REGION Network 14: I42.5 - Tank Vent Valve 2 Feedback Closed (CV-441-B)
   // True = CLOSED, False = NOT
   RUNG wire#powerrail
      Contact( "Tank 4S Tank Vent Valve 2 Feedback - Closed" )
      Coil( "20_TANKS_IP_DATA".RIO_04.SECOND_TANK.TANK_VENT_B_CLSD )
   END_RUNG
   // the same network as SCL:
   "20_TANKS_IP_DATA".RIO_04.SECOND_TANK.TANK_VENT_B_CLSD := "Tank 4S Tank Vent Valve 2 Feedback - Closed";
END_REGION

REGION Network 15: I42.6 - Spare Input Destination Accesed from Warning FC
   // True = N/A, False = N/A
END_REGION

REGION Network 16: I42.7 - Spare Input
   // True = N/A, False = N/A
   RUNG wire#powerrail
      Contact( "RIO4_SPR_DI_142_7" )
      Coil( "20_TANKS_IP_DATA".RIO_04.SECOND_TANK.SPARE_DI_7 )
   END_RUNG
   // the same network as SCL:
   "20_TANKS_IP_DATA".RIO_04.SECOND_TANK.SPARE_DI_7 := "RIO4_SPR_DI_142_7";
END_REGION

REGION Network 17: I45.0 - Tank Level HIHI - (LS-425) - First Tank
   // True = OK, False = HIHI
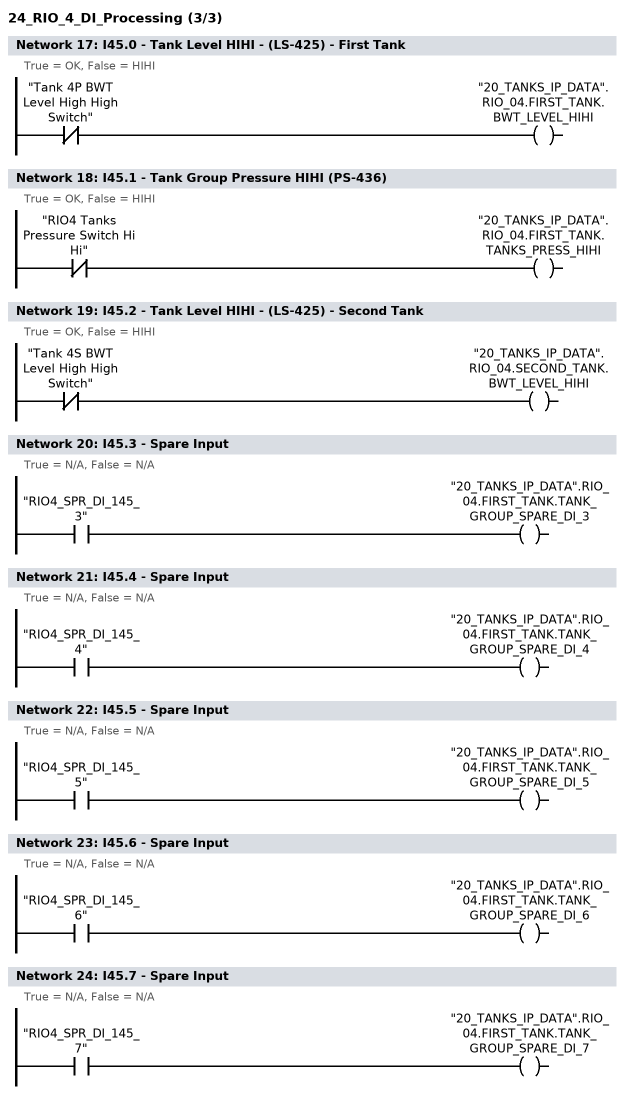
   RUNG wire#powerrail
      I_Contact( "Tank 4P BWT Level High High Switch" )
      Coil( "20_TANKS_IP_DATA".RIO_04.FIRST_TANK.BWT_LEVEL_HIHI )
   END_RUNG
   // the same network as SCL:
   "20_TANKS_IP_DATA".RIO_04.FIRST_TANK.BWT_LEVEL_HIHI := NOT "Tank 4P BWT Level High High Switch";
END_REGION

REGION Network 18: I45.1 - Tank Group Pressure HIHI (PS-436)
   // True = OK, False = HIHI
   RUNG wire#powerrail
      I_Contact( "RIO4 Tanks Pressure Switch Hi Hi" )
      Coil( "20_TANKS_IP_DATA".RIO_04.FIRST_TANK.TANKS_PRESS_HIHI )
   END_RUNG
   // the same network as SCL:
   "20_TANKS_IP_DATA".RIO_04.FIRST_TANK.TANKS_PRESS_HIHI := NOT "RIO4 Tanks Pressure Switch Hi Hi";
END_REGION

REGION Network 19: I45.2 - Tank Level HIHI - (LS-425) - Second Tank
   // True = OK, False = HIHI
   RUNG wire#powerrail
      I_Contact( "Tank 4S BWT Level High High Switch" )
      Coil( "20_TANKS_IP_DATA".RIO_04.SECOND_TANK.BWT_LEVEL_HIHI )
   END_RUNG
   // the same network as SCL:
   "20_TANKS_IP_DATA".RIO_04.SECOND_TANK.BWT_LEVEL_HIHI := NOT "Tank 4S BWT Level High High Switch";
END_REGION

REGION Network 20: I45.3 - Spare Input
   // True = N/A, False = N/A
   RUNG wire#powerrail
      Contact( "RIO4_SPR_DI_145_3" )
      Coil( "20_TANKS_IP_DATA".RIO_04.FIRST_TANK.TANK_GROUP_SPARE_DI_3 )
   END_RUNG
   // the same network as SCL:
   "20_TANKS_IP_DATA".RIO_04.FIRST_TANK.TANK_GROUP_SPARE_DI_3 := "RIO4_SPR_DI_145_3";
END_REGION

REGION Network 21: I45.4 - Spare Input
   // True = N/A, False = N/A
   RUNG wire#powerrail
      Contact( "RIO4_SPR_DI_145_4" )
      Coil( "20_TANKS_IP_DATA".RIO_04.FIRST_TANK.TANK_GROUP_SPARE_DI_4 )
   END_RUNG
   // the same network as SCL:
   "20_TANKS_IP_DATA".RIO_04.FIRST_TANK.TANK_GROUP_SPARE_DI_4 := "RIO4_SPR_DI_145_4";
END_REGION

REGION Network 22: I45.5 - Spare Input
   // True = N/A, False = N/A
   RUNG wire#powerrail
      Contact( "RIO4_SPR_DI_145_5" )
      Coil( "20_TANKS_IP_DATA".RIO_04.FIRST_TANK.TANK_GROUP_SPARE_DI_5 )
   END_RUNG
   // the same network as SCL:
   "20_TANKS_IP_DATA".RIO_04.FIRST_TANK.TANK_GROUP_SPARE_DI_5 := "RIO4_SPR_DI_145_5";
END_REGION

REGION Network 23: I45.6 - Spare Input
   // True = N/A, False = N/A
   RUNG wire#powerrail
      Contact( "RIO4_SPR_DI_145_6" )
      Coil( "20_TANKS_IP_DATA".RIO_04.FIRST_TANK.TANK_GROUP_SPARE_DI_6 )
   END_RUNG
   // the same network as SCL:
   "20_TANKS_IP_DATA".RIO_04.FIRST_TANK.TANK_GROUP_SPARE_DI_6 := "RIO4_SPR_DI_145_6";
END_REGION

REGION Network 24: I45.7 - Spare Input
   // True = N/A, False = N/A
   RUNG wire#powerrail
      Contact( "RIO4_SPR_DI_145_7" )
      Coil( "20_TANKS_IP_DATA".RIO_04.FIRST_TANK.TANK_GROUP_SPARE_DI_7 )
   END_RUNG
   // the same network as SCL:
   "20_TANKS_IP_DATA".RIO_04.FIRST_TANK.TANK_GROUP_SPARE_DI_7 := "RIO4_SPR_DI_145_7";
END_REGION
END_FUNCTION

FUNCTION "25_RIO_5_DI_Processing" : Void   // FC25, LAD
TITLE = RIO Rack Digital Input Processing (Tank 1 = 5P, Tank 2 = 5S)
{ S7_Optimized_Access := 'TRUE' }
AUTHOR : JRS
VERSION : 0.1
// To process raw inputs prior to code use
BEGIN

REGION Network 1: I51.0 - Gas To Tank Valve Feedback Open (CV-422)
   // True = OPEN, False = NOT
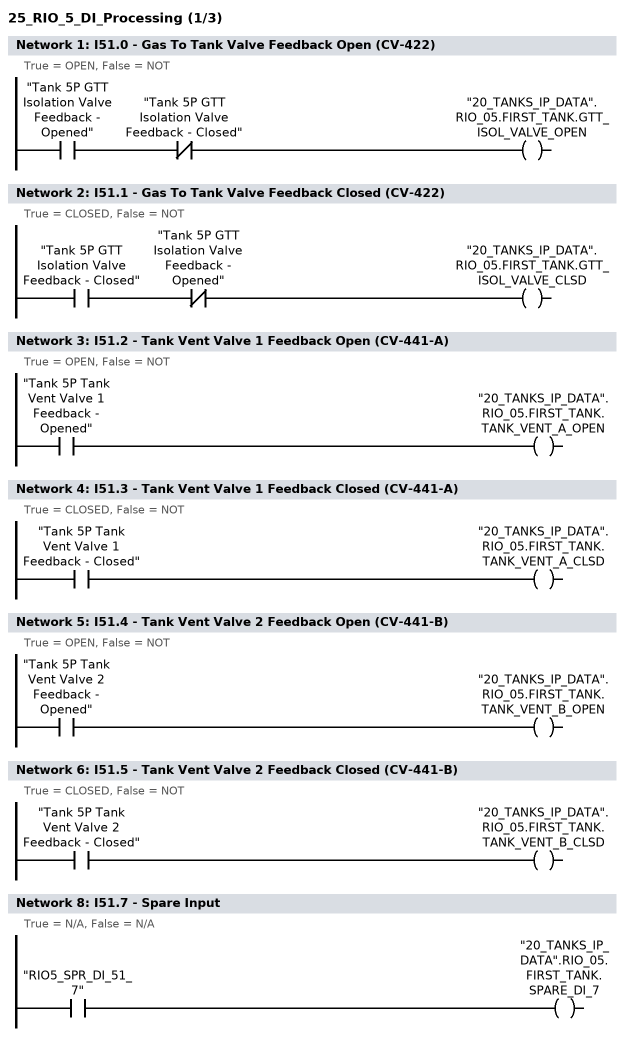
   RUNG wire#powerrail
      Contact( "Tank 5P GTT Isolation Valve Feedback - Opened" )
      I_Contact( "Tank 5P GTT Isolation Valve Feedback - Closed" )
      Coil( "20_TANKS_IP_DATA".RIO_05.FIRST_TANK.GTT_ISOL_VALVE_OPEN )
   END_RUNG
   // the same network as SCL:
   "20_TANKS_IP_DATA".RIO_05.FIRST_TANK.GTT_ISOL_VALVE_OPEN := "Tank 5P GTT Isolation Valve Feedback - Opened" AND NOT "Tank 5P GTT Isolation Valve Feedback - Closed";
END_REGION

REGION Network 2: I51.1 - Gas To Tank Valve Feedback Closed (CV-422)
   // True = CLOSED, False = NOT
   RUNG wire#powerrail
      Contact( "Tank 5P GTT Isolation Valve Feedback - Closed" )
      I_Contact( "Tank 5P GTT Isolation Valve Feedback - Opened" )
      Coil( "20_TANKS_IP_DATA".RIO_05.FIRST_TANK.GTT_ISOL_VALVE_CLSD )
   END_RUNG
   // the same network as SCL:
   "20_TANKS_IP_DATA".RIO_05.FIRST_TANK.GTT_ISOL_VALVE_CLSD := "Tank 5P GTT Isolation Valve Feedback - Closed" AND NOT "Tank 5P GTT Isolation Valve Feedback - Opened";
END_REGION

REGION Network 3: I51.2 - Tank Vent Valve 1 Feedback Open (CV-441-A)
   // True = OPEN, False = NOT
   RUNG wire#powerrail
      Contact( "Tank 5P Tank Vent Valve 1 Feedback - Opened" )
      Coil( "20_TANKS_IP_DATA".RIO_05.FIRST_TANK.TANK_VENT_A_OPEN )
   END_RUNG
   // the same network as SCL:
   "20_TANKS_IP_DATA".RIO_05.FIRST_TANK.TANK_VENT_A_OPEN := "Tank 5P Tank Vent Valve 1 Feedback - Opened";
END_REGION

REGION Network 4: I51.3 - Tank Vent Valve 1 Feedback Closed (CV-441-A)
   // True = CLOSED, False = NOT
   RUNG wire#powerrail
      Contact( "Tank 5P Tank Vent Valve 1 Feedback - Closed" )
      Coil( "20_TANKS_IP_DATA".RIO_05.FIRST_TANK.TANK_VENT_A_CLSD )
   END_RUNG
   // the same network as SCL:
   "20_TANKS_IP_DATA".RIO_05.FIRST_TANK.TANK_VENT_A_CLSD := "Tank 5P Tank Vent Valve 1 Feedback - Closed";
END_REGION

REGION Network 5: I51.4 - Tank Vent Valve 2 Feedback Open (CV-441-B)
   // True = OPEN, False = NOT
   RUNG wire#powerrail
      Contact( "Tank 5P Tank Vent Valve 2 Feedback - Opened" )
      Coil( "20_TANKS_IP_DATA".RIO_05.FIRST_TANK.TANK_VENT_B_OPEN )
   END_RUNG
   // the same network as SCL:
   "20_TANKS_IP_DATA".RIO_05.FIRST_TANK.TANK_VENT_B_OPEN := "Tank 5P Tank Vent Valve 2 Feedback - Opened";
END_REGION

REGION Network 6: I51.5 - Tank Vent Valve 2 Feedback Closed (CV-441-B)
   // True = CLOSED, False = NOT
   RUNG wire#powerrail
      Contact( "Tank 5P Tank Vent Valve 2 Feedback - Closed" )
      Coil( "20_TANKS_IP_DATA".RIO_05.FIRST_TANK.TANK_VENT_B_CLSD )
   END_RUNG
   // the same network as SCL:
   "20_TANKS_IP_DATA".RIO_05.FIRST_TANK.TANK_VENT_B_CLSD := "Tank 5P Tank Vent Valve 2 Feedback - Closed";
END_REGION

REGION Network 7: I51.6 - Spare Input Destination Accesed from Warning FC
   // True = N/A, False = N/A
END_REGION

REGION Network 8: I51.7 - Spare Input
   // True = N/A, False = N/A
   RUNG wire#powerrail
      Contact( "RIO5_SPR_DI_51_7" )
      Coil( "20_TANKS_IP_DATA".RIO_05.FIRST_TANK.SPARE_DI_7 )
   END_RUNG
   // the same network as SCL:
   "20_TANKS_IP_DATA".RIO_05.FIRST_TANK.SPARE_DI_7 := "RIO5_SPR_DI_51_7";
END_REGION

REGION Network 9: I54.0 - Gas To Tank Valve Feedback Open (CV-422)
   // True = OPEN, False = NOT
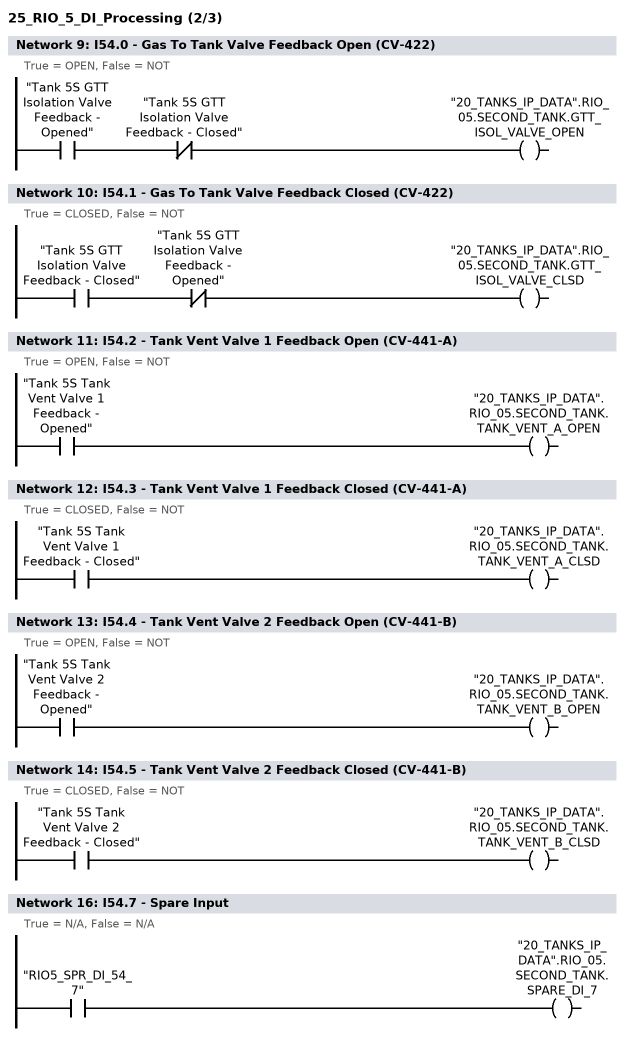
   RUNG wire#powerrail
      Contact( "Tank 5S GTT Isolation Valve Feedback - Opened" )
      I_Contact( "Tank 5S GTT Isolation Valve Feedback - Closed" )
      Coil( "20_TANKS_IP_DATA".RIO_05.SECOND_TANK.GTT_ISOL_VALVE_OPEN )
   END_RUNG
   // the same network as SCL:
   "20_TANKS_IP_DATA".RIO_05.SECOND_TANK.GTT_ISOL_VALVE_OPEN := "Tank 5S GTT Isolation Valve Feedback - Opened" AND NOT "Tank 5S GTT Isolation Valve Feedback - Closed";
END_REGION

REGION Network 10: I54.1 - Gas To Tank Valve Feedback Closed (CV-422)
   // True = CLOSED, False = NOT
   RUNG wire#powerrail
      Contact( "Tank 5S GTT Isolation Valve Feedback - Closed" )
      I_Contact( "Tank 5S GTT Isolation Valve Feedback - Opened" )
      Coil( "20_TANKS_IP_DATA".RIO_05.SECOND_TANK.GTT_ISOL_VALVE_CLSD )
   END_RUNG
   // the same network as SCL:
   "20_TANKS_IP_DATA".RIO_05.SECOND_TANK.GTT_ISOL_VALVE_CLSD := "Tank 5S GTT Isolation Valve Feedback - Closed" AND NOT "Tank 5S GTT Isolation Valve Feedback - Opened";
END_REGION

REGION Network 11: I54.2 - Tank Vent Valve 1 Feedback Open (CV-441-A)
   // True = OPEN, False = NOT
   RUNG wire#powerrail
      Contact( "Tank 5S Tank Vent Valve 1 Feedback - Opened" )
      Coil( "20_TANKS_IP_DATA".RIO_05.SECOND_TANK.TANK_VENT_A_OPEN )
   END_RUNG
   // the same network as SCL:
   "20_TANKS_IP_DATA".RIO_05.SECOND_TANK.TANK_VENT_A_OPEN := "Tank 5S Tank Vent Valve 1 Feedback - Opened";
END_REGION

REGION Network 12: I54.3 - Tank Vent Valve 1 Feedback Closed (CV-441-A)
   // True = CLOSED, False = NOT
   RUNG wire#powerrail
      Contact( "Tank 5S Tank Vent Valve 1 Feedback - Closed" )
      Coil( "20_TANKS_IP_DATA".RIO_05.SECOND_TANK.TANK_VENT_A_CLSD )
   END_RUNG
   // the same network as SCL:
   "20_TANKS_IP_DATA".RIO_05.SECOND_TANK.TANK_VENT_A_CLSD := "Tank 5S Tank Vent Valve 1 Feedback - Closed";
END_REGION

REGION Network 13: I54.4 - Tank Vent Valve 2 Feedback Open (CV-441-B)
   // True = OPEN, False = NOT
   RUNG wire#powerrail
      Contact( "Tank 5S Tank Vent Valve 2 Feedback - Opened" )
      Coil( "20_TANKS_IP_DATA".RIO_05.SECOND_TANK.TANK_VENT_B_OPEN )
   END_RUNG
   // the same network as SCL:
   "20_TANKS_IP_DATA".RIO_05.SECOND_TANK.TANK_VENT_B_OPEN := "Tank 5S Tank Vent Valve 2 Feedback - Opened";
END_REGION

REGION Network 14: I54.5 - Tank Vent Valve 2 Feedback Closed (CV-441-B)
   // True = CLOSED, False = NOT
   RUNG wire#powerrail
      Contact( "Tank 5S Tank Vent Valve 2 Feedback - Closed" )
      Coil( "20_TANKS_IP_DATA".RIO_05.SECOND_TANK.TANK_VENT_B_CLSD )
   END_RUNG
   // the same network as SCL:
   "20_TANKS_IP_DATA".RIO_05.SECOND_TANK.TANK_VENT_B_CLSD := "Tank 5S Tank Vent Valve 2 Feedback - Closed";
END_REGION

REGION Network 15: I54.6 - Spare Input Destination Accesed from Warning FC
   // True = N/A, False = N/A
END_REGION

REGION Network 16: I54.7 - Spare Input
   // True = N/A, False = N/A
   RUNG wire#powerrail
      Contact( "RIO5_SPR_DI_54_7" )
      Coil( "20_TANKS_IP_DATA".RIO_05.SECOND_TANK.SPARE_DI_7 )
   END_RUNG
   // the same network as SCL:
   "20_TANKS_IP_DATA".RIO_05.SECOND_TANK.SPARE_DI_7 := "RIO5_SPR_DI_54_7";
END_REGION

REGION Network 17: I57.0 - Tank Level HIHI - (LS-425) - First Tank
   // True = OK, False = HIHI
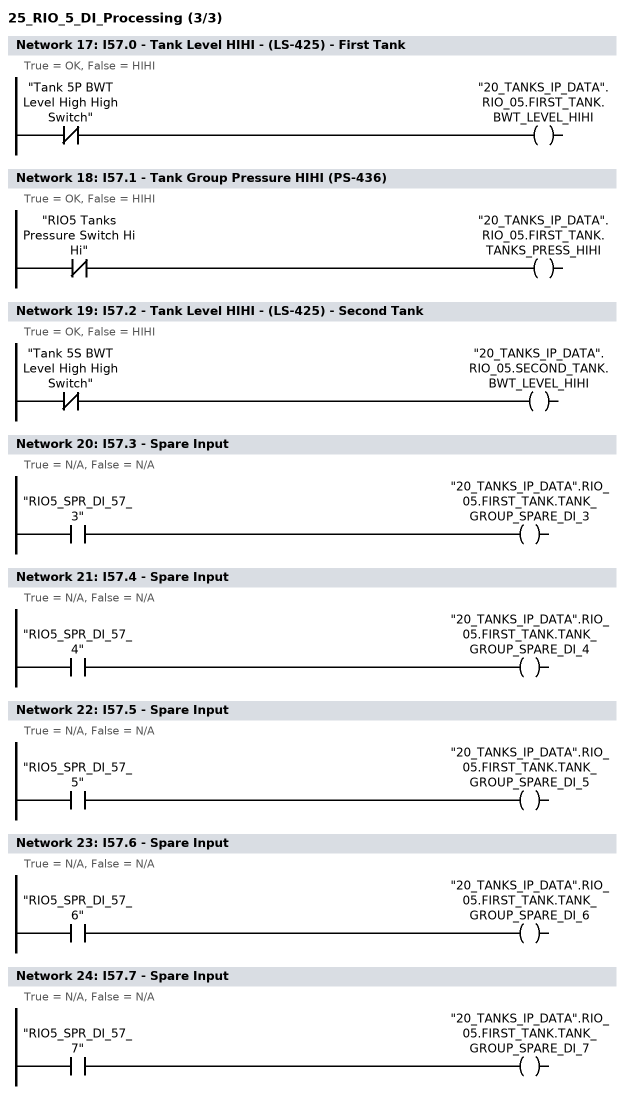
   RUNG wire#powerrail
      I_Contact( "Tank 5P BWT Level High High Switch" )
      Coil( "20_TANKS_IP_DATA".RIO_05.FIRST_TANK.BWT_LEVEL_HIHI )
   END_RUNG
   // the same network as SCL:
   "20_TANKS_IP_DATA".RIO_05.FIRST_TANK.BWT_LEVEL_HIHI := NOT "Tank 5P BWT Level High High Switch";
END_REGION

REGION Network 18: I57.1 - Tank Group Pressure HIHI (PS-436)
   // True = OK, False = HIHI
   RUNG wire#powerrail
      I_Contact( "RIO5 Tanks Pressure Switch Hi Hi" )
      Coil( "20_TANKS_IP_DATA".RIO_05.FIRST_TANK.TANKS_PRESS_HIHI )
   END_RUNG
   // the same network as SCL:
   "20_TANKS_IP_DATA".RIO_05.FIRST_TANK.TANKS_PRESS_HIHI := NOT "RIO5 Tanks Pressure Switch Hi Hi";
END_REGION

REGION Network 19: I57.2 - Tank Level HIHI - (LS-425) - Second Tank
   // True = OK, False = HIHI
   RUNG wire#powerrail
      I_Contact( "Tank 5S BWT Level High High Switch" )
      Coil( "20_TANKS_IP_DATA".RIO_05.SECOND_TANK.BWT_LEVEL_HIHI )
   END_RUNG
   // the same network as SCL:
   "20_TANKS_IP_DATA".RIO_05.SECOND_TANK.BWT_LEVEL_HIHI := NOT "Tank 5S BWT Level High High Switch";
END_REGION

REGION Network 20: I57.3 - Spare Input
   // True = N/A, False = N/A
   RUNG wire#powerrail
      Contact( "RIO5_SPR_DI_57_3" )
      Coil( "20_TANKS_IP_DATA".RIO_05.FIRST_TANK.TANK_GROUP_SPARE_DI_3 )
   END_RUNG
   // the same network as SCL:
   "20_TANKS_IP_DATA".RIO_05.FIRST_TANK.TANK_GROUP_SPARE_DI_3 := "RIO5_SPR_DI_57_3";
END_REGION

REGION Network 21: I57.4 - Spare Input
   // True = N/A, False = N/A
   RUNG wire#powerrail
      Contact( "RIO5_SPR_DI_57_4" )
      Coil( "20_TANKS_IP_DATA".RIO_05.FIRST_TANK.TANK_GROUP_SPARE_DI_4 )
   END_RUNG
   // the same network as SCL:
   "20_TANKS_IP_DATA".RIO_05.FIRST_TANK.TANK_GROUP_SPARE_DI_4 := "RIO5_SPR_DI_57_4";
END_REGION

REGION Network 22: I57.5 - Spare Input
   // True = N/A, False = N/A
   RUNG wire#powerrail
      Contact( "RIO5_SPR_DI_57_5" )
      Coil( "20_TANKS_IP_DATA".RIO_05.FIRST_TANK.TANK_GROUP_SPARE_DI_5 )
   END_RUNG
   // the same network as SCL:
   "20_TANKS_IP_DATA".RIO_05.FIRST_TANK.TANK_GROUP_SPARE_DI_5 := "RIO5_SPR_DI_57_5";
END_REGION

REGION Network 23: I57.6 - Spare Input
   // True = N/A, False = N/A
   RUNG wire#powerrail
      Contact( "RIO5_SPR_DI_57_6" )
      Coil( "20_TANKS_IP_DATA".RIO_05.FIRST_TANK.TANK_GROUP_SPARE_DI_6 )
   END_RUNG
   // the same network as SCL:
   "20_TANKS_IP_DATA".RIO_05.FIRST_TANK.TANK_GROUP_SPARE_DI_6 := "RIO5_SPR_DI_57_6";
END_REGION

REGION Network 24: I57.7 - Spare Input
   // True = N/A, False = N/A
   RUNG wire#powerrail
      Contact( "RIO5_SPR_DI_57_7" )
      Coil( "20_TANKS_IP_DATA".RIO_05.FIRST_TANK.TANK_GROUP_SPARE_DI_7 )
   END_RUNG
   // the same network as SCL:
   "20_TANKS_IP_DATA".RIO_05.FIRST_TANK.TANK_GROUP_SPARE_DI_7 := "RIO5_SPR_DI_57_7";
END_REGION
END_FUNCTION

FUNCTION "26_RIO_6_DI_Processing" : Void   // FC26, LAD
TITLE = RIO Rack Digital Input Processing (Tank 1 = 6P, Tank 2 = 6S)
{ S7_Optimized_Access := 'TRUE' }
AUTHOR : JRS
VERSION : 0.1
// To process raw inputs prior to code use
BEGIN

REGION Network 1: I60.0 - Gas To Tank Valve Feedback Open (CV-422)
   // True = OPEN, False = NOT
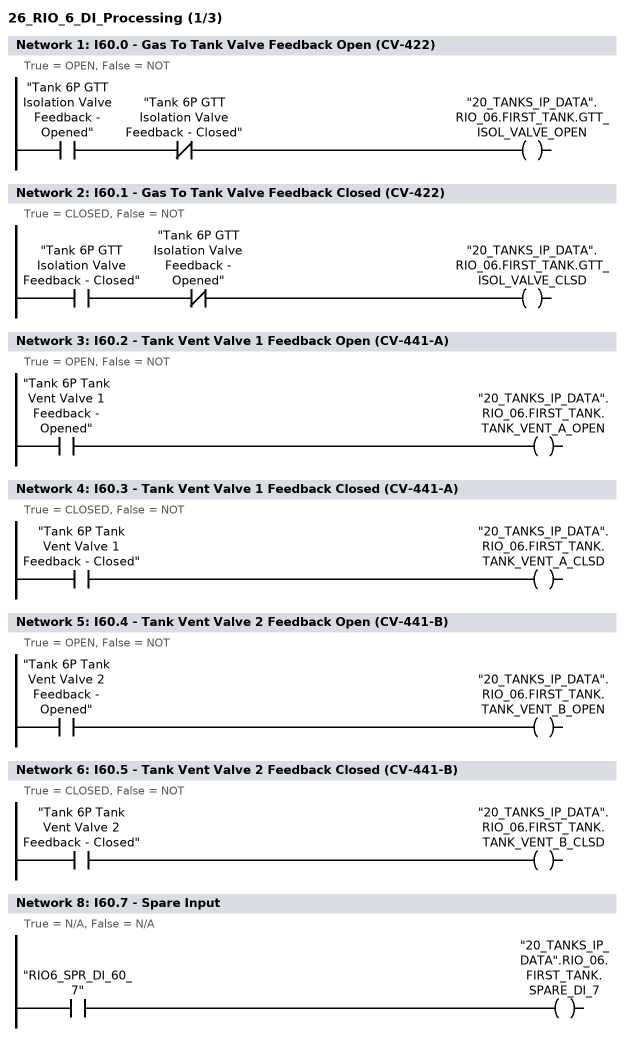
   RUNG wire#powerrail
      Contact( "Tank 6P GTT Isolation Valve Feedback - Opened" )
      I_Contact( "Tank 6P GTT Isolation Valve Feedback - Closed" )
      Coil( "20_TANKS_IP_DATA".RIO_06.FIRST_TANK.GTT_ISOL_VALVE_OPEN )
   END_RUNG
   // the same network as SCL:
   "20_TANKS_IP_DATA".RIO_06.FIRST_TANK.GTT_ISOL_VALVE_OPEN := "Tank 6P GTT Isolation Valve Feedback - Opened" AND NOT "Tank 6P GTT Isolation Valve Feedback - Closed";
END_REGION

REGION Network 2: I60.1 - Gas To Tank Valve Feedback Closed (CV-422)
   // True = CLOSED, False = NOT
   RUNG wire#powerrail
      Contact( "Tank 6P GTT Isolation Valve Feedback - Closed" )
      I_Contact( "Tank 6P GTT Isolation Valve Feedback - Opened" )
      Coil( "20_TANKS_IP_DATA".RIO_06.FIRST_TANK.GTT_ISOL_VALVE_CLSD )
   END_RUNG
   // the same network as SCL:
   "20_TANKS_IP_DATA".RIO_06.FIRST_TANK.GTT_ISOL_VALVE_CLSD := "Tank 6P GTT Isolation Valve Feedback - Closed" AND NOT "Tank 6P GTT Isolation Valve Feedback - Opened";
END_REGION

REGION Network 3: I60.2 - Tank Vent Valve 1 Feedback Open (CV-441-A)
   // True = OPEN, False = NOT
   RUNG wire#powerrail
      Contact( "Tank 6P Tank Vent Valve 1 Feedback - Opened" )
      Coil( "20_TANKS_IP_DATA".RIO_06.FIRST_TANK.TANK_VENT_A_OPEN )
   END_RUNG
   // the same network as SCL:
   "20_TANKS_IP_DATA".RIO_06.FIRST_TANK.TANK_VENT_A_OPEN := "Tank 6P Tank Vent Valve 1 Feedback - Opened";
END_REGION

REGION Network 4: I60.3 - Tank Vent Valve 1 Feedback Closed (CV-441-A)
   // True = CLOSED, False = NOT
   RUNG wire#powerrail
      Contact( "Tank 6P Tank Vent Valve 1 Feedback - Closed" )
      Coil( "20_TANKS_IP_DATA".RIO_06.FIRST_TANK.TANK_VENT_A_CLSD )
   END_RUNG
   // the same network as SCL:
   "20_TANKS_IP_DATA".RIO_06.FIRST_TANK.TANK_VENT_A_CLSD := "Tank 6P Tank Vent Valve 1 Feedback - Closed";
END_REGION

REGION Network 5: I60.4 - Tank Vent Valve 2 Feedback Open (CV-441-B)
   // True = OPEN, False = NOT
   RUNG wire#powerrail
      Contact( "Tank 6P Tank Vent Valve 2 Feedback - Opened" )
      Coil( "20_TANKS_IP_DATA".RIO_06.FIRST_TANK.TANK_VENT_B_OPEN )
   END_RUNG
   // the same network as SCL:
   "20_TANKS_IP_DATA".RIO_06.FIRST_TANK.TANK_VENT_B_OPEN := "Tank 6P Tank Vent Valve 2 Feedback - Opened";
END_REGION

REGION Network 6: I60.5 - Tank Vent Valve 2 Feedback Closed (CV-441-B)
   // True = CLOSED, False = NOT
   RUNG wire#powerrail
      Contact( "Tank 6P Tank Vent Valve 2 Feedback - Closed" )
      Coil( "20_TANKS_IP_DATA".RIO_06.FIRST_TANK.TANK_VENT_B_CLSD )
   END_RUNG
   // the same network as SCL:
   "20_TANKS_IP_DATA".RIO_06.FIRST_TANK.TANK_VENT_B_CLSD := "Tank 6P Tank Vent Valve 2 Feedback - Closed";
END_REGION

REGION Network 7: I60.6 - Spare Input Destination Accesed from Warning FC
   // True = N/A, False = N/A
END_REGION

REGION Network 8: I60.7 - Spare Input
   // True = N/A, False = N/A
   RUNG wire#powerrail
      Contact( "RIO6_SPR_DI_60_7" )
      Coil( "20_TANKS_IP_DATA".RIO_06.FIRST_TANK.SPARE_DI_7 )
   END_RUNG
   // the same network as SCL:
   "20_TANKS_IP_DATA".RIO_06.FIRST_TANK.SPARE_DI_7 := "RIO6_SPR_DI_60_7";
END_REGION

REGION Network 9: I63.0 - Gas To Tank Valve Feedback Open (CV-422)
   // True = OPEN, False = NOT
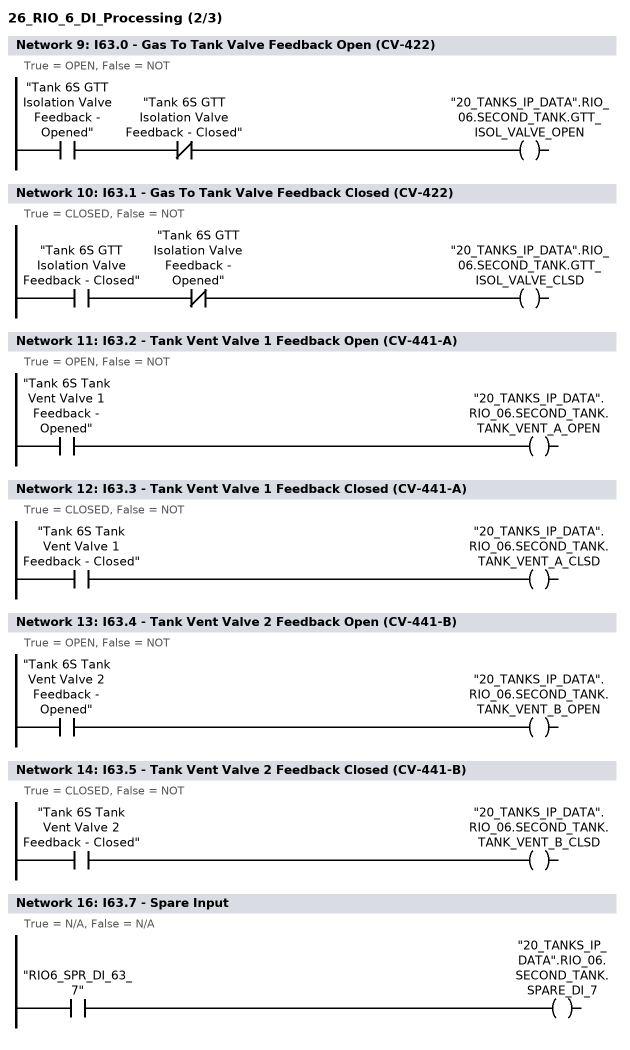
   RUNG wire#powerrail
      Contact( "Tank 6S GTT Isolation Valve Feedback - Opened" )
      I_Contact( "Tank 6S GTT Isolation Valve Feedback - Closed" )
      Coil( "20_TANKS_IP_DATA".RIO_06.SECOND_TANK.GTT_ISOL_VALVE_OPEN )
   END_RUNG
   // the same network as SCL:
   "20_TANKS_IP_DATA".RIO_06.SECOND_TANK.GTT_ISOL_VALVE_OPEN := "Tank 6S GTT Isolation Valve Feedback - Opened" AND NOT "Tank 6S GTT Isolation Valve Feedback - Closed";
END_REGION

REGION Network 10: I63.1 - Gas To Tank Valve Feedback Closed (CV-422)
   // True = CLOSED, False = NOT
   RUNG wire#powerrail
      Contact( "Tank 6S GTT Isolation Valve Feedback - Closed" )
      I_Contact( "Tank 6S GTT Isolation Valve Feedback - Opened" )
      Coil( "20_TANKS_IP_DATA".RIO_06.SECOND_TANK.GTT_ISOL_VALVE_CLSD )
   END_RUNG
   // the same network as SCL:
   "20_TANKS_IP_DATA".RIO_06.SECOND_TANK.GTT_ISOL_VALVE_CLSD := "Tank 6S GTT Isolation Valve Feedback - Closed" AND NOT "Tank 6S GTT Isolation Valve Feedback - Opened";
END_REGION

REGION Network 11: I63.2 - Tank Vent Valve 1 Feedback Open (CV-441-A)
   // True = OPEN, False = NOT
   RUNG wire#powerrail
      Contact( "Tank 6S Tank Vent Valve 1 Feedback - Opened" )
      Coil( "20_TANKS_IP_DATA".RIO_06.SECOND_TANK.TANK_VENT_A_OPEN )
   END_RUNG
   // the same network as SCL:
   "20_TANKS_IP_DATA".RIO_06.SECOND_TANK.TANK_VENT_A_OPEN := "Tank 6S Tank Vent Valve 1 Feedback - Opened";
END_REGION

REGION Network 12: I63.3 - Tank Vent Valve 1 Feedback Closed (CV-441-A)
   // True = CLOSED, False = NOT
   RUNG wire#powerrail
      Contact( "Tank 6S Tank Vent Valve 1 Feedback - Closed" )
      Coil( "20_TANKS_IP_DATA".RIO_06.SECOND_TANK.TANK_VENT_A_CLSD )
   END_RUNG
   // the same network as SCL:
   "20_TANKS_IP_DATA".RIO_06.SECOND_TANK.TANK_VENT_A_CLSD := "Tank 6S Tank Vent Valve 1 Feedback - Closed";
END_REGION

REGION Network 13: I63.4 - Tank Vent Valve 2 Feedback Open (CV-441-B)
   // True = OPEN, False = NOT
   RUNG wire#powerrail
      Contact( "Tank 6S Tank Vent Valve 2 Feedback - Opened" )
      Coil( "20_TANKS_IP_DATA".RIO_06.SECOND_TANK.TANK_VENT_B_OPEN )
   END_RUNG
   // the same network as SCL:
   "20_TANKS_IP_DATA".RIO_06.SECOND_TANK.TANK_VENT_B_OPEN := "Tank 6S Tank Vent Valve 2 Feedback - Opened";
END_REGION

REGION Network 14: I63.5 - Tank Vent Valve 2 Feedback Closed (CV-441-B)
   // True = CLOSED, False = NOT
   RUNG wire#powerrail
      Contact( "Tank 6S Tank Vent Valve 2 Feedback - Closed" )
      Coil( "20_TANKS_IP_DATA".RIO_06.SECOND_TANK.TANK_VENT_B_CLSD )
   END_RUNG
   // the same network as SCL:
   "20_TANKS_IP_DATA".RIO_06.SECOND_TANK.TANK_VENT_B_CLSD := "Tank 6S Tank Vent Valve 2 Feedback - Closed";
END_REGION

REGION Network 15: I63.6 - Spare Input Destination Accesed from Warning FC
   // True = N/A, False = N/A
END_REGION

REGION Network 16: I63.7 - Spare Input
   // True = N/A, False = N/A
   RUNG wire#powerrail
      Contact( "RIO6_SPR_DI_63_7" )
      Coil( "20_TANKS_IP_DATA".RIO_06.SECOND_TANK.SPARE_DI_7 )
   END_RUNG
   // the same network as SCL:
   "20_TANKS_IP_DATA".RIO_06.SECOND_TANK.SPARE_DI_7 := "RIO6_SPR_DI_63_7";
END_REGION

REGION Network 17: I66.0 - Tank Level HIHI - (LS-425) - First Tank
   // True = OK, False = HIHI
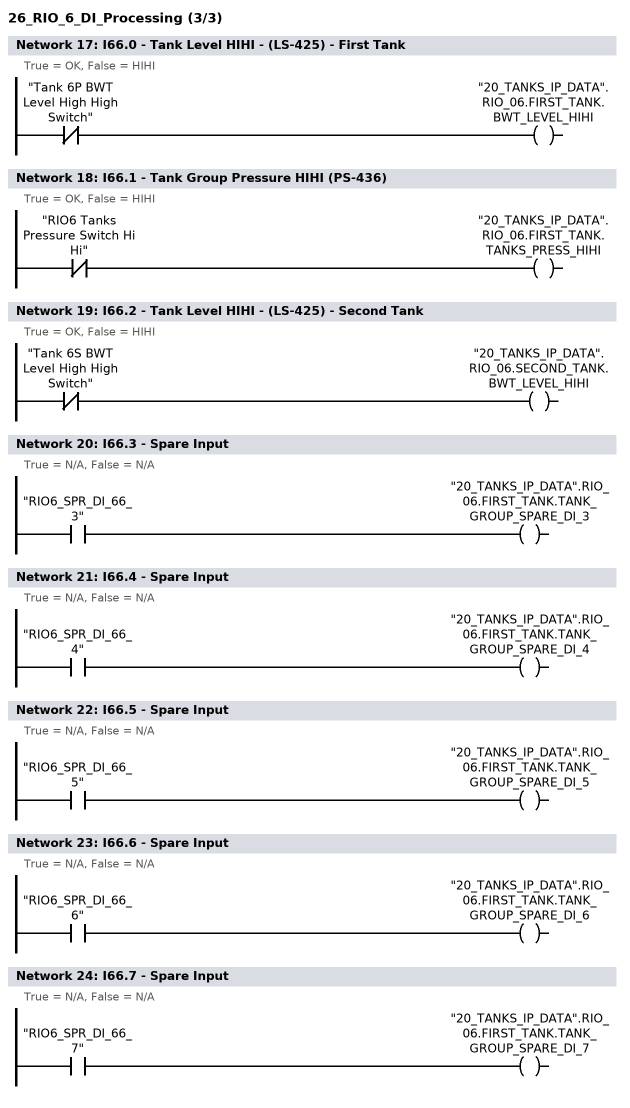
   RUNG wire#powerrail
      I_Contact( "Tank 6P BWT Level High High Switch" )
      Coil( "20_TANKS_IP_DATA".RIO_06.FIRST_TANK.BWT_LEVEL_HIHI )
   END_RUNG
   // the same network as SCL:
   "20_TANKS_IP_DATA".RIO_06.FIRST_TANK.BWT_LEVEL_HIHI := NOT "Tank 6P BWT Level High High Switch";
END_REGION

REGION Network 18: I66.1 - Tank Group Pressure HIHI (PS-436)
   // True = OK, False = HIHI
   RUNG wire#powerrail
      I_Contact( "RIO6 Tanks Pressure Switch Hi Hi" )
      Coil( "20_TANKS_IP_DATA".RIO_06.FIRST_TANK.TANKS_PRESS_HIHI )
   END_RUNG
   // the same network as SCL:
   "20_TANKS_IP_DATA".RIO_06.FIRST_TANK.TANKS_PRESS_HIHI := NOT "RIO6 Tanks Pressure Switch Hi Hi";
END_REGION

REGION Network 19: I66.2 - Tank Level HIHI - (LS-425) - Second Tank
   // True = OK, False = HIHI
   RUNG wire#powerrail
      I_Contact( "Tank 6S BWT Level High High Switch" )
      Coil( "20_TANKS_IP_DATA".RIO_06.SECOND_TANK.BWT_LEVEL_HIHI )
   END_RUNG
   // the same network as SCL:
   "20_TANKS_IP_DATA".RIO_06.SECOND_TANK.BWT_LEVEL_HIHI := NOT "Tank 6S BWT Level High High Switch";
END_REGION

REGION Network 20: I66.3 - Spare Input
   // True = N/A, False = N/A
   RUNG wire#powerrail
      Contact( "RIO6_SPR_DI_66_3" )
      Coil( "20_TANKS_IP_DATA".RIO_06.FIRST_TANK.TANK_GROUP_SPARE_DI_3 )
   END_RUNG
   // the same network as SCL:
   "20_TANKS_IP_DATA".RIO_06.FIRST_TANK.TANK_GROUP_SPARE_DI_3 := "RIO6_SPR_DI_66_3";
END_REGION

REGION Network 21: I66.4 - Spare Input
   // True = N/A, False = N/A
   RUNG wire#powerrail
      Contact( "RIO6_SPR_DI_66_4" )
      Coil( "20_TANKS_IP_DATA".RIO_06.FIRST_TANK.TANK_GROUP_SPARE_DI_4 )
   END_RUNG
   // the same network as SCL:
   "20_TANKS_IP_DATA".RIO_06.FIRST_TANK.TANK_GROUP_SPARE_DI_4 := "RIO6_SPR_DI_66_4";
END_REGION

REGION Network 22: I66.5 - Spare Input
   // True = N/A, False = N/A
   RUNG wire#powerrail
      Contact( "RIO6_SPR_DI_66_5" )
      Coil( "20_TANKS_IP_DATA".RIO_06.FIRST_TANK.TANK_GROUP_SPARE_DI_5 )
   END_RUNG
   // the same network as SCL:
   "20_TANKS_IP_DATA".RIO_06.FIRST_TANK.TANK_GROUP_SPARE_DI_5 := "RIO6_SPR_DI_66_5";
END_REGION

REGION Network 23: I66.6 - Spare Input
   // True = N/A, False = N/A
   RUNG wire#powerrail
      Contact( "RIO6_SPR_DI_66_6" )
      Coil( "20_TANKS_IP_DATA".RIO_06.FIRST_TANK.TANK_GROUP_SPARE_DI_6 )
   END_RUNG
   // the same network as SCL:
   "20_TANKS_IP_DATA".RIO_06.FIRST_TANK.TANK_GROUP_SPARE_DI_6 := "RIO6_SPR_DI_66_6";
END_REGION

REGION Network 24: I66.7 - Spare Input
   // True = N/A, False = N/A
   RUNG wire#powerrail
      Contact( "RIO6_SPR_DI_66_7" )
      Coil( "20_TANKS_IP_DATA".RIO_06.FIRST_TANK.TANK_GROUP_SPARE_DI_7 )
   END_RUNG
   // the same network as SCL:
   "20_TANKS_IP_DATA".RIO_06.FIRST_TANK.TANK_GROUP_SPARE_DI_7 := "RIO6_SPR_DI_66_7";
END_REGION
END_FUNCTION

FUNCTION "27_RIO_7_DI_Processing" : Void   // FC27, LAD
TITLE = RIO Rack Digital Input Processing (Tank 1 = APT)
{ S7_Optimized_Access := 'TRUE' }
AUTHOR : JRS
VERSION : 0.1
// To process raw inputs prior to code use
BEGIN

REGION Network 1: I75.0 - Gas To Tank Valve Feedback Open (CV-422)
   // True = OPEN, False = NOT
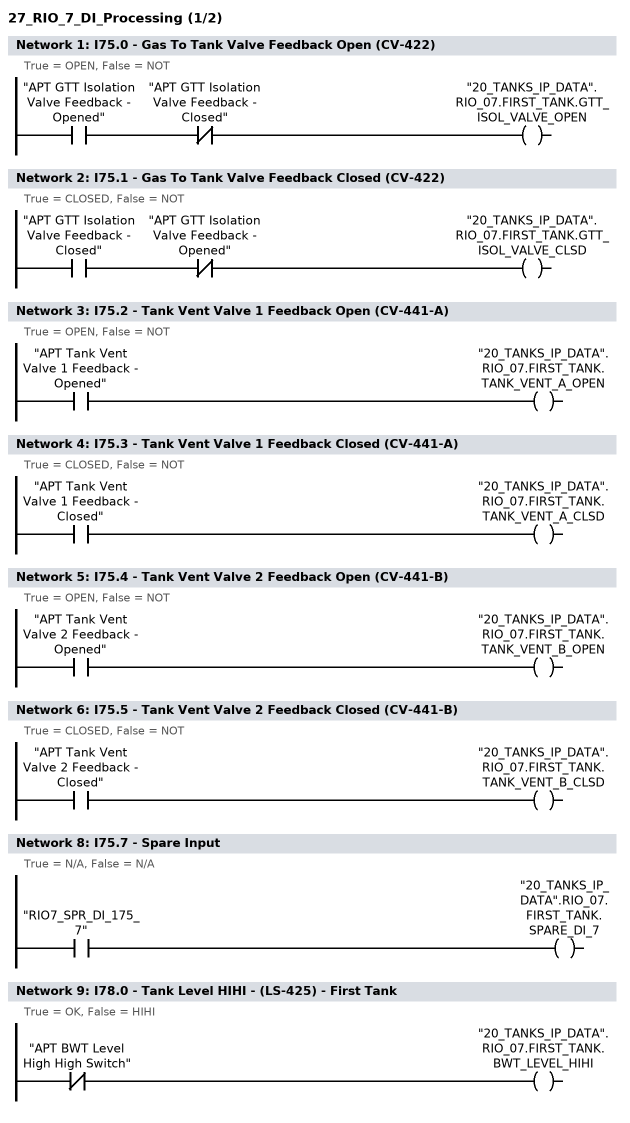
   RUNG wire#powerrail
      Contact( "APT GTT Isolation Valve Feedback - Opened" )
      I_Contact( "APT GTT Isolation Valve Feedback - Closed" )
      Coil( "20_TANKS_IP_DATA".RIO_07.FIRST_TANK.GTT_ISOL_VALVE_OPEN )
   END_RUNG
   // the same network as SCL:
   "20_TANKS_IP_DATA".RIO_07.FIRST_TANK.GTT_ISOL_VALVE_OPEN := "APT GTT Isolation Valve Feedback - Opened" AND NOT "APT GTT Isolation Valve Feedback - Closed";
END_REGION

REGION Network 2: I75.1 - Gas To Tank Valve Feedback Closed (CV-422)
   // True = CLOSED, False = NOT
   RUNG wire#powerrail
      Contact( "APT GTT Isolation Valve Feedback - Closed" )
      I_Contact( "APT GTT Isolation Valve Feedback - Opened" )
      Coil( "20_TANKS_IP_DATA".RIO_07.FIRST_TANK.GTT_ISOL_VALVE_CLSD )
   END_RUNG
   // the same network as SCL:
   "20_TANKS_IP_DATA".RIO_07.FIRST_TANK.GTT_ISOL_VALVE_CLSD := "APT GTT Isolation Valve Feedback - Closed" AND NOT "APT GTT Isolation Valve Feedback - Opened";
END_REGION
